   1709: 'Spare_Fault_1709', class No Acknowledgement, trigger "DB302_HMI_Faults_Carrier26_Faults_2" bit 12
   1710: 'Spare_Fault_1710', class No Acknowledgement, trigger "DB302_HMI_Faults_Carrier26_Faults_2" bit 13
   1711: 'Spare_Fault_1711', class No Acknowledgement, trigger "DB302_HMI_Faults_Carrier26_Faults_2" bit 14
   1712: 'Spare_Fault_1712', class No Acknowledgement, trigger "DB302_HMI_Faults_Carrier26_Faults_2" bit 15
   1713: 'Spare_Fault_1713', class No Acknowledgement, trigger "DB302_HMI_Faults_Carrier26_Faults_3" bit 0
   1714: 'Spare_Fault_1714', class No Acknowledgement, trigger "DB302_HMI_Faults_Carrier26_Faults_3" bit 1
   1715: 'Spare_Fault_1715', class No Acknowledgement, trigger "DB302_HMI_Faults_Carrier26_Faults_3" bit 2
   1716: 'Spare_Fault_1716', class No Acknowledgement, trigger "DB302_HMI_Faults_Carrier26_Faults_3" bit 3
   1717: 'Spare_Fault_1717', class No Acknowledgement, trigger "DB302_HMI_Faults_Carrier26_Faults_3" bit 4
   1718: 'Spare_Fault_1718', class No Acknowledgement, trigger "DB302_HMI_Faults_Carrier26_Faults_3" bit 5
   1719: 'Spare_Fault_1719', class No Acknowledgement, trigger "DB302_HMI_Faults_Carrier26_Faults_3" bit 6
   1720: 'Spare_Fault_1720', class No Acknowledgement, trigger "DB302_HMI_Faults_Carrier26_Faults_3" bit 7
   1721: 'Spare_Fault_1721', class No Acknowledgement, trigger "DB302_HMI_Faults_Carrier26_Faults_3" bit 8
   1722: 'Spare_Fault_1722', class No Acknowledgement, trigger "DB302_HMI_Faults_Carrier26_Faults_3" bit 9
   1723: 'Spare_Fault_1723', class No Acknowledgement, trigger "DB302_HMI_Faults_Carrier26_Faults_3" bit 10
   1724: 'Spare_Fault_1724', class No Acknowledgement, trigger "DB302_HMI_Faults_Carrier26_Faults_3" bit 11
   1725: 'Spare_Fault_1725', class No Acknowledgement, trigger "DB302_HMI_Faults_Carrier26_Faults_3" bit 12
   1726: 'Spare_Fault_1726', class No Acknowledgement, trigger "DB302_HMI_Faults_Carrier26_Faults_3" bit 13
   1727: 'Spare_Fault_1727', class No Acknowledgement, trigger "DB302_HMI_Faults_Carrier26_Faults_3" bit 14
   1728: 'Spare_Fault_1728', class No Acknowledgement, trigger "DB302_HMI_Faults_Carrier26_Faults_3" bit 15
   1729: 'Carrier 27 Disconnect Open Power Fault DI11.0', class No Acknowledgement, trigger "DB302_HMI_Faults_Carrier27_Faults_0" bit 0
   1730: 'Carrier 27 Drive Profinet Comm Fault', class No Acknowledgement, trigger "DB302_HMI_Faults_Carrier27_Faults_0" bit 1
   1731: 'Carrier 27 Production Stop Not Reset', class No Acknowledgement, trigger "DB302_HMI_Faults_Carrier27_Faults_0" bit 2
   1732: 'Carrier 27 CB02122 Tripped', class No Acknowledgement, trigger "DB302_HMI_Faults_Carrier27_Faults_0" bit 3
   1733: 'Carrier 27 CB02123 Tripped', class No Acknowledgement, trigger "DB302_HMI_Faults_Carrier27_Faults_0" bit 4
   1734: 'Carrier 27 AUX1 CB Tripped', class No Acknowledgement, trigger "DB302_HMI_Faults_Carrier27_Faults_0" bit 5
   1735: 'Carrier 27 AUX2 CB Tripped', class No Acknowledgement, trigger "DB302_HMI_Faults_Carrier27_Faults_0" bit 6
   1736: 'Carrier 27 PLC Not Communicating', class No Acknowledgement, trigger "DB302_HMI_Faults_Carrier27_Faults_0" bit 7
   1737: 'Carrier 27 Safe Input Card Fault', class No Acknowledgement, trigger "DB302_HMI_Faults_Carrier27_Faults_0" bit 8
   1738: 'Carrier 27 Safe Output Card Fault', class No Acknowledgement, trigger "DB302_HMI_Faults_Carrier27_Faults_0" bit 9
   1739: 'Carrier 27 Standard Input Card Fault', class No Acknowledgement, trigger "DB302_HMI_Faults_Carrier27_Faults_0" bit 10
   1740: 'Carrier 27 Standard Output Card Fault', class No Acknowledgement, trigger "DB302_HMI_Faults_Carrier27_Faults_0" bit 11
   1741: 'Carrier 27 Encoder Position Fault', class No Acknowledgement, trigger "DB302_HMI_Faults_Carrier27_Faults_0" bit 12
   1742: 'Carrier 27 Encoder Internal Error', class No Acknowledgement, trigger "DB302_HMI_Faults_Carrier27_Faults_0" bit 13
   1743: 'Carrier 27 Encoder Comm Fault', class No Acknowledgement, trigger "DB302_HMI_Faults_Carrier27_Faults_0" bit 14
   1744: 'Carrier 27 HMI Comm Fault', class No Acknowledgement, trigger "DB302_HMI_Faults_Carrier27_Faults_0" bit 15
   1745: 'Carrier 27 Crash Detection Fault', class No Acknowledgement, trigger "DB302_HMI_Faults_Carrier27_Faults_1" bit 0
   1746: 'Carrier 27 Carrier Number Invalid', class No Acknowledgement, trigger "DB302_HMI_Faults_Carrier27_Faults_1" bit 1
   1747: 'Carrier 27 Drive: PROFINET configuration error', class No Acknowledgement, trigger "DB302_HMI_Faults_Carrier27_Faults_1" bit 2
   1748: 'Carrier 27 Drive: Error internal communications', class No Acknowledgement, trigger "DB302_HMI_Faults_Carrier27_Faults_1" bit 3
   1749: 'Carrier 27 Drive: Motor overtemperature', class No Acknowledgement, trigger "DB302_HMI_Faults_Carrier27_Faults_1" bit 4
   1750: 'Carrier 27 Drive: Motor overcurrent', class No Acknowledgement, trigger "DB302_HMI_Faults_Carrier27_Faults_1" bit 5
   1751: 'Carrier 27 Drive: Infeed or power unit not ready', class No Acknowledgement, trigger "DB302_HMI_Faults_Carrier27_Faults_1" bit 6
   1752: 'Carrier 27 Drive: Short-circuit/ground fault detected', class No Acknowledgement, trigger "DB302_HMI_Faults_Carrier27_Faults_1" bit 7
   1753: 'Carrier 27 Drive: PROFINET Setpoint timeout', class No Acknowledgement, trigger "DB302_HMI_Faults_Carrier27_Faults_1" bit 8
   1754: 'Carrier 27 Power unit: Overcurrent', class No Acknowledgement, trigger "DB302_HMI_Faults_Carrier27_Faults_1" bit 9
   1755: 'Carrier 27 Power unit: DC link voltage overvoltage', class No Acknowledgement, trigger "DB302_HMI_Faults_Carrier27_Faults_1" bit 10
   1756: 'Carrier 27 Power unit: DC link voltage undervoltage', class No Acknowledgement, trigger "DB302_HMI_Faults_Carrier27_Faults_1" bit 11
   1757: 'Carrier 27 Power unit: Line phase failure in main circuit', class No Acknowledgement, trigger "DB302_HMI_Faults_Carrier27_Faults_1" bit 12
   1758: 'Carrier 27 Power unit: Phase failure motor cable', class No Acknowledgement, trigger "DB302_HMI_Faults_Carrier27_Faults_1" bit 13
   1759: 'Carrier 27 Power unit: Ground fault', class No Acknowledgement, trigger "DB302_HMI_Faults_Carrier27_Faults_1" bit 14
   1760: 'Spare_Fault_1760', class No Acknowledgement, trigger "DB302_HMI_Faults_Carrier27_Faults_1" bit 15
   1761: 'Carrier 27 Motion Off Fault', class No Acknowledgement, trigger "DB302_HMI_Faults_Carrier27_Faults_2" bit 0
   1762: 'Carrier 27 Motion On Fault', class No Acknowledgement, trigger "DB302_HMI_Faults_Carrier27_Faults_2" bit 1
   1763: 'Carrier 27 Spacing Fault', class No Acknowledgement, trigger "DB302_HMI_Faults_Carrier27_Faults_2" bit 2
   1764: 'Carrier 27 Duplicate Carrier Number Fault', class No Acknowledgement, trigger "DB302_HMI_Faults_Carrier27_Faults_2" bit 3
   1765: 'Spare_Fault_1765', class No Acknowledgement, trigger "DB302_HMI_Faults_Carrier27_Faults_2" bit 4
   1766: 'Spare_Fault_1766', class No Acknowledgement, trigger "DB302_HMI_Faults_Carrier27_Faults_2" bit 5
   1767: 'Spare_Fault_1767', class No Acknowledgement, trigger "DB302_HMI_Faults_Carrier27_Faults_2" bit 6
   1768: 'Spare_Fault_1768', class No Acknowledgement, trigger "DB302_HMI_Faults_Carrier27_Faults_2" bit 7
   1769: 'Spare_Fault_1769', class No Acknowledgement, trigger "DB302_HMI_Faults_Carrier27_Faults_2" bit 8
   1770: 'Spare_Fault_1770', class No Acknowledgement, trigger "DB302_HMI_Faults_Carrier27_Faults_2" bit 9
   1771: 'Spare_Fault_1771', class No Acknowledgement, trigger "DB302_HMI_Faults_Carrier27_Faults_2" bit 10
   1772: 'Spare_Fault_1772', class No Acknowledgement, trigger "DB302_HMI_Faults_Carrier27_Faults_2" bit 11
   1773: 'Spare_Fault_1773', class No Acknowledgement, trigger "DB302_HMI_Faults_Carrier27_Faults_2" bit 12
   1774: 'Spare_Fault_1774', class No Acknowledgement, trigger "DB302_HMI_Faults_Carrier27_Faults_2" bit 13
   1775: 'Spare_Fault_1775', class No Acknowledgement, trigger "DB302_HMI_Faults_Carrier27_Faults_2" bit 14
   1776: 'Spare_Fault_1776', class No Acknowledgement, trigger "DB302_HMI_Faults_Carrier27_Faults_2" bit 15
   1777: 'Spare_Fault_1777', class No Acknowledgement, trigger "DB302_HMI_Faults_Carrier27_Faults_3" bit 0
   1778: 'Spare_Fault_1778', class No Acknowledgement, trigger "DB302_HMI_Faults_Carrier27_Faults_3" bit 1
   1779: 'Spare_Fault_1779', class No Acknowledgement, trigger "DB302_HMI_Faults_Carrier27_Faults_3" bit 2
   1780: 'Spare_Fault_1780', class No Acknowledgement, trigger "DB302_HMI_Faults_Carrier27_Faults_3" bit 3
   1781: 'Spare_Fault_1781', class No Acknowledgement, trigger "DB302_HMI_Faults_Carrier27_Faults_3" bit 4
   1782: 'Spare_Fault_1782', class No Acknowledgement, trigger "DB302_HMI_Faults_Carrier27_Faults_3" bit 5
   1783: 'Spare_Fault_1783', class No Acknowledgement, trigger "DB302_HMI_Faults_Carrier27_Faults_3" bit 6
   1784: 'Spare_Fault_1784', class No Acknowledgement, trigger "DB302_HMI_Faults_Carrier27_Faults_3" bit 7
   1785: 'Spare_Fault_1785', class No Acknowledgement, trigger "DB302_HMI_Faults_Carrier27_Faults_3" bit 8
   1786: 'Spare_Fault_1786', class No Acknowledgement, trigger "DB302_HMI_Faults_Carrier27_Faults_3" bit 9
   1787: 'Spare_Fault_1787', class No Acknowledgement, trigger "DB302_HMI_Faults_Carrier27_Faults_3" bit 10
   1788: 'Spare_Fault_1788', class No Acknowledgement, trigger "DB302_HMI_Faults_Carrier27_Faults_3" bit 11
   1789: 'Spare_Fault_1789', class No Acknowledgement, trigger "DB302_HMI_Faults_Carrier27_Faults_3" bit 12
   1790: 'Spare_Fault_1790', class No Acknowledgement, trigger "DB302_HMI_Faults_Carrier27_Faults_3" bit 13
   1791: 'Spare_Fault_1791', class No Acknowledgement, trigger "DB302_HMI_Faults_Carrier27_Faults_3" bit 14
   1792: 'Spare_Fault_1792', class No Acknowledgement, trigger "DB302_HMI_Faults_Carrier27_Faults_3" bit 15
   1793: 'Carrier 28 Disconnect Open Power Fault DI11.0', class No Acknowledgement, trigger "DB302_HMI_Faults_Carrier28_Faults_0" bit 0
   1794: 'Carrier 28 Drive Profinet Comm Fault', class No Acknowledgement, trigger "DB302_HMI_Faults_Carrier28_Faults_0" bit 1
   1795: 'Carrier 28 Production Stop Not Reset', class No Acknowledgement, trigger "DB302_HMI_Faults_Carrier28_Faults_0" bit 2
   1796: 'Carrier 28 CB02122 Tripped', class No Acknowledgement, trigger "DB302_HMI_Faults_Carrier28_Faults_0" bit 3
   1797: 'Carrier 28 CB02123 Tripped', class No Acknowledgement, trigger "DB302_HMI_Faults_Carrier28_Faults_0" bit 4
   1798: 'Carrier 28 AUX1 CB Tripped', class No Acknowledgement, trigger "DB302_HMI_Faults_Carrier28_Faults_0" bit 5
   1799: 'Carrier 28 AUX2 CB Tripped', class No Acknowledgement, trigger "DB302_HMI_Faults_Carrier28_Faults_0" bit 6
   1800: 'Carrier 28 PLC Not Communicating', class No Acknowledgement, trigger "DB302_HMI_Faults_Carrier28_Faults_0" bit 7
   1801: 'Carrier 28 Safe Input Card Fault', class No Acknowledgement, trigger "DB302_HMI_Faults_Carrier28_Faults_0" bit 8
   1802: 'Carrier 28 Safe Output Card Fault', class No Acknowledgement, trigger "DB302_HMI_Faults_Carrier28_Faults_0" bit 9
   1803: 'Carrier 28 Standard Input Card Fault', class No Acknowledgement, trigger "DB302_HMI_Faults_Carrier28_Faults_0" bit 10
   1804: 'Carrier 28 Standard Output Card Fault', class No Acknowledgement, trigger "DB302_HMI_Faults_Carrier28_Faults_0" bit 11
   1805: 'Carrier 28 Encoder Position Fault', class No Acknowledgement, trigger "DB302_HMI_Faults_Carrier28_Faults_0" bit 12
   1806: 'Carrier 28 Encoder Internal Error', class No Acknowledgement, trigger "DB302_HMI_Faults_Carrier28_Faults_0" bit 13
   1807: 'Carrier 28 Encoder Comm Fault', class No Acknowledgement, trigger "DB302_HMI_Faults_Carrier28_Faults_0" bit 14
   1808: 'Carrier 28 HMI Comm Fault', class No Acknowledgement, trigger "DB302_HMI_Faults_Carrier28_Faults_0" bit 15
   1809: 'Carrier 28 Crash Detection Fault', class No Acknowledgement, trigger "DB302_HMI_Faults_Carrier28_Faults_1" bit 0
   1810: 'Carrier 28 Carrier Number Invalid', class No Acknowledgement, trigger "DB302_HMI_Faults_Carrier28_Faults_1" bit 1
   1811: 'Carrier 28 Drive: PROFINET configuration error', class No Acknowledgement, trigger "DB302_HMI_Faults_Carrier28_Faults_1" bit 2
   1812: 'Carrier 28 Drive: Error internal communications', class No Acknowledgement, trigger "DB302_HMI_Faults_Carrier28_Faults_1" bit 3
   1813: 'Carrier 28 Drive: Motor overtemperature', class No Acknowledgement, trigger "DB302_HMI_Faults_Carrier28_Faults_1" bit 4
   1814: 'Carrier 28 Drive: Motor overcurrent', class No Acknowledgement, trigger "DB302_HMI_Faults_Carrier28_Faults_1" bit 5
   1815: 'Carrier 28 Drive: Infeed or power unit not ready', class No Acknowledgement, trigger "DB302_HMI_Faults_Carrier28_Faults_1" bit 6
   1816: 'Carrier 28 Drive: Short-circuit/ground fault detected', class No Acknowledgement, trigger "DB302_HMI_Faults_Carrier28_Faults_1" bit 7
   1817: 'Carrier 28 Drive: PROFINET Setpoint timeout', class No Acknowledgement, trigger "DB302_HMI_Faults_Carrier28_Faults_1" bit 8
   1818: 'Carrier 28 Power unit: Overcurrent', class No Acknowledgement, trigger "DB302_HMI_Faults_Carrier28_Faults_1" bit 9
   1819: 'Carrier 28 Power unit: DC link voltage overvoltage', class No Acknowledgement, trigger "DB302_HMI_Faults_Carrier28_Faults_1" bit 10
   1820: 'Carrier 28 Power unit: DC link voltage undervoltage', class No Acknowledgement, trigger "DB302_HMI_Faults_Carrier28_Faults_1" bit 11
   1821: 'Carrier 28 Power unit: Line phase failure in main circuit', class No Acknowledgement, trigger "DB302_HMI_Faults_Carrier28_Faults_1" bit 12
   1822: 'Carrier 28 Power unit: Phase failure motor cable', class No Acknowledgement, trigger "DB302_HMI_Faults_Carrier28_Faults_1" bit 13
   1823: 'Carrier 28 Power unit: Ground fault', class No Acknowledgement, trigger "DB302_HMI_Faults_Carrier28_Faults_1" bit 14
   1824: 'Spare_Fault_1824', class No Acknowledgement, trigger "DB302_HMI_Faults_Carrier28_Faults_1" bit 15
   1825: 'Carrier 28 Motion Off Fault', class No Acknowledgement, trigger "DB302_HMI_Faults_Carrier28_Faults_2" bit 0
   1826: 'Carrier 28 Motion On Fault', class No Acknowledgement, trigger "DB302_HMI_Faults_Carrier28_Faults_2" bit 1
   1827: 'Carrier 28 Spacing Fault', class No Acknowledgement, trigger "DB302_HMI_Faults_Carrier28_Faults_2" bit 2
   1828: 'Carrier 28 Duplicate Carrier Number Fault', class No Acknowledgement, trigger "DB302_HMI_Faults_Carrier28_Faults_2" bit 3
   1829: 'Spare_Fault_1829', class No Acknowledgement, trigger "DB302_HMI_Faults_Carrier28_Faults_2" bit 4
   1830: 'Spare_Fault_1830', class No Acknowledgement, trigger "DB302_HMI_Faults_Carrier28_Faults_2" bit 5
   1831: 'Spare_Fault_1831', class No Acknowledgement, trigger "DB302_HMI_Faults_Carrier28_Faults_2" bit 6
   1832: 'Spare_Fault_1832', class No Acknowledgement, trigger "DB302_HMI_Faults_Carrier28_Faults_2" bit 7
   1833: 'Spare_Fault_1833', class No Acknowledgement, trigger "DB302_HMI_Faults_Carrier28_Faults_2" bit 8
   1834: 'Spare_Fault_1834', class No Acknowledgement, trigger "DB302_HMI_Faults_Carrier28_Faults_2" bit 9
   1835: 'Spare_Fault_1835', class No Acknowledgement, trigger "DB302_HMI_Faults_Carrier28_Faults_2" bit 10
   1836: 'Spare_Fault_1836', class No Acknowledgement, trigger "DB302_HMI_Faults_Carrier28_Faults_2" bit 11
   1837: 'Spare_Fault_1837', class No Acknowledgement, trigger "DB302_HMI_Faults_Carrier28_Faults_2" bit 12
   1838: 'Spare_Fault_1838', class No Acknowledgement, trigger "DB302_HMI_Faults_Carrier28_Faults_2" bit 13
   1839: 'Spare_Fault_1839', class No Acknowledgement, trigger "DB302_HMI_Faults_Carrier28_Faults_2" bit 14
   1840: 'Spare_Fault_1840', class No Acknowledgement, trigger "DB302_HMI_Faults_Carrier28_Faults_2" bit 15
   1841: 'Spare_Fault_1841', class No Acknowledgement, trigger "DB302_HMI_Faults_Carrier28_Faults_3" bit 0
   1842: 'Spare_Fault_1842', class No Acknowledgement, trigger "DB302_HMI_Faults_Carrier28_Faults_3" bit 1
   1843: 'Spare_Fault_1843', class No Acknowledgement, trigger "DB302_HMI_Faults_Carrier28_Faults_3" bit 2
   1844: 'Spare_Fault_1844', class No Acknowledgement, trigger "DB302_HMI_Faults_Carrier28_Faults_3" bit 3
   1845: 'Spare_Fault_1845', class No Acknowledgement, trigger "DB302_HMI_Faults_Carrier28_Faults_3" bit 4
   1846: 'Spare_Fault_1846', class No Acknowledgement, trigger "DB302_HMI_Faults_Carrier28_Faults_3" bit 5
   1847: 'Spare_Fault_1847', class No Acknowledgement, trigger "DB302_HMI_Faults_Carrier28_Faults_3" bit 6
   1848: 'Spare_Fault_1848', class No Acknowledgement, trigger "DB302_HMI_Faults_Carrier28_Faults_3" bit 7
   1849: 'Spare_Fault_1849', class No Acknowledgement, trigger "DB302_HMI_Faults_Carrier28_Faults_3" bit 8
   1850: 'Spare_Fault_1850', class No Acknowledgement, trigger "DB302_HMI_Faults_Carrier28_Faults_3" bit 9
   1851: 'Spare_Fault_1851', class No Acknowledgement, trigger "DB302_HMI_Faults_Carrier28_Faults_3" bit 10
   1852: 'Spare_Fault_1852', class No Acknowledgement, trigger "DB302_HMI_Faults_Carrier28_Faults_3" bit 11
   1853: 'Spare_Fault_1853', class No Acknowledgement, trigger "DB302_HMI_Faults_Carrier28_Faults_3" bit 12
   1854: 'Spare_Fault_1854', class No Acknowledgement, trigger "DB302_HMI_Faults_Carrier28_Faults_3" bit 13
   1855: 'Spare_Fault_1855', class No Acknowledgement, trigger "DB302_HMI_Faults_Carrier28_Faults_3" bit 14
   1856: 'Spare_Fault_1856', class No Acknowledgement, trigger "DB302_HMI_Faults_Carrier28_Faults_3" bit 15
   1857: 'Carrier 29 Disconnect Open Power Fault DI11.0', class No Acknowledgement, trigger "DB302_HMI_Faults_Carrier29_Faults_0" bit 0
   1858: 'Carrier 29 Drive Profinet Comm Fault', class No Acknowledgement, trigger "DB302_HMI_Faults_Carrier29_Faults_0" bit 1
   1859: 'Carrier 29 Production Stop Not Reset', class No Acknowledgement, trigger "DB302_HMI_Faults_Carrier29_Faults_0" bit 2
   1860: 'Carrier 29 CB02122 Tripped', class No Acknowledgement, trigger "DB302_HMI_Faults_Carrier29_Faults_0" bit 3
   1861: 'Carrier 29 CB02123 Tripped', class No Acknowledgement, trigger "DB302_HMI_Faults_Carrier29_Faults_0" bit 4
   1862: 'Carrier 29 AUX1 CB Tripped', class No Acknowledgement, trigger "DB302_HMI_Faults_Carrier29_Faults_0" bit 5
   1863: 'Carrier 29 AUX2 CB Tripped', class No Acknowledgement, trigger "DB302_HMI_Faults_Carrier29_Faults_0" bit 6
   1864: 'Carrier 29 PLC Not Communicating', class No Acknowledgement, trigger "DB302_HMI_Faults_Carrier29_Faults_0" bit 7
   1865: 'Carrier 29 Safe Input Card Fault', class No Acknowledgement, trigger "DB302_HMI_Faults_Carrier29_Faults_0" bit 8
   1866: 'Carrier 29 Safe Output Card Fault', class No Acknowledgement, trigger "DB302_HMI_Faults_Carrier29_Faults_0" bit 9
   1867: 'Carrier 29 Standard Input Card Fault', class No Acknowledgement, trigger "DB302_HMI_Faults_Carrier29_Faults_0" bit 10
   1868: 'Carrier 29 Standard Output Card Fault', class No Acknowledgement, trigger "DB302_HMI_Faults_Carrier29_Faults_0" bit 11
   1869: 'Carrier 29 Encoder Position Fault', class No Acknowledgement, trigger "DB302_HMI_Faults_Carrier29_Faults_0" bit 12
   1870: 'Carrier 29 Encoder Internal Error', class No Acknowledgement, trigger "DB302_HMI_Faults_Carrier29_Faults_0" bit 13
   1871: 'Carrier 29 Encoder Comm Fault', class No Acknowledgement, trigger "DB302_HMI_Faults_Carrier29_Faults_0" bit 14
   1872: 'Carrier 29 HMI Comm Fault', class No Acknowledgement, trigger "DB302_HMI_Faults_Carrier29_Faults_0" bit 15
   1873: 'Carrier 29 Crash Detection Fault', class No Acknowledgement, trigger "DB302_HMI_Faults_Carrier29_Faults_1" bit 0
   1874: 'Carrier 29 Carrier Number Invalid', class No Acknowledgement, trigger "DB302_HMI_Faults_Carrier29_Faults_1" bit 1
   1875: 'Carrier 29 Drive: PROFINET configuration error', class No Acknowledgement, trigger "DB302_HMI_Faults_Carrier29_Faults_1" bit 2
   1876: 'Carrier 29 Drive: Error internal communications', class No Acknowledgement, trigger "DB302_HMI_Faults_Carrier29_Faults_1" bit 3
   1877: 'Carrier 29 Drive: Motor overtemperature', class No Acknowledgement, trigger "DB302_HMI_Faults_Carrier29_Faults_1" bit 4
   1878: 'Carrier 29 Drive: Motor overcurrent', class No Acknowledgement, trigger "DB302_HMI_Faults_Carrier29_Faults_1" bit 5
   1879: 'Carrier 29 Drive: Infeed or power unit not ready', class No Acknowledgement, trigger "DB302_HMI_Faults_Carrier29_Faults_1" bit 6
   1880: 'Carrier 29 Drive: Short-circuit/ground fault detected', class No Acknowledgement, trigger "DB302_HMI_Faults_Carrier29_Faults_1" bit 7
   1881: 'Carrier 29 Drive: PROFINET Setpoint timeout', class No Acknowledgement, trigger "DB302_HMI_Faults_Carrier29_Faults_1" bit 8
   1882: 'Carrier 29 Power unit: Overcurrent', class No Acknowledgement, trigger "DB302_HMI_Faults_Carrier29_Faults_1" bit 9
   1883: 'Carrier 29 Power unit: DC link voltage overvoltage', class No Acknowledgement, trigger "DB302_HMI_Faults_Carrier29_Faults_1" bit 10
   1884: 'Carrier 29 Power unit: DC link voltage undervoltage', class No Acknowledgement, trigger "DB302_HMI_Faults_Carrier29_Faults_1" bit 11
   1885: 'Carrier 29 Power unit: Line phase failure in main circuit', class No Acknowledgement, trigger "DB302_HMI_Faults_Carrier29_Faults_1" bit 12
   1886: 'Carrier 29 Power unit: Phase failure motor cable', class No Acknowledgement, trigger "DB302_HMI_Faults_Carrier29_Faults_1" bit 13
   1887: 'Carrier 29 Power unit: Ground fault', class No Acknowledgement, trigger "DB302_HMI_Faults_Carrier29_Faults_1" bit 14
   1888: 'Spare_Fault_1888', class No Acknowledgement, trigger "DB302_HMI_Faults_Carrier29_Faults_1" bit 15
   1889: 'Carrier 29 Motion Off Fault', class No Acknowledgement, trigger "DB302_HMI_Faults_Carrier29_Faults_2" bit 0
   1890: 'Carrier 29 Motion On Fault', class No Acknowledgement, trigger "DB302_HMI_Faults_Carrier29_Faults_2" bit 1
   1891: 'Carrier 29 Spacing Fault', class No Acknowledgement, trigger "DB302_HMI_Faults_Carrier29_Faults_2" bit 2
   1892: 'Carrier 29 Duplicate Carrier Number Fault', class No Acknowledgement, trigger "DB302_HMI_Faults_Carrier29_Faults_2" bit 3
   1893: 'Spare_Fault_1893', class No Acknowledgement, trigger "DB302_HMI_Faults_Carrier29_Faults_2" bit 4
   1894: 'Spare_Fault_1894', class No Acknowledgement, trigger "DB302_HMI_Faults_Carrier29_Faults_2" bit 5
   1895: 'Spare_Fault_1895', class No Acknowledgement, trigger "DB302_HMI_Faults_Carrier29_Faults_2" bit 6
   1896: 'Spare_Fault_1896', class No Acknowledgement, trigger "DB302_HMI_Faults_Carrier29_Faults_2" bit 7
   1897: 'Spare_Fault_1897', class No Acknowledgement, trigger "DB302_HMI_Faults_Carrier29_Faults_2" bit 8
   1898: 'Spare_Fault_1898', class No Acknowledgement, trigger "DB302_HMI_Faults_Carrier29_Faults_2" bit 9
   1899: 'Spare_Fault_1899', class No Acknowledgement, trigger "DB302_HMI_Faults_Carrier29_Faults_2" bit 10
   1900: 'Spare_Fault_1900', class No Acknowledgement, trigger "DB302_HMI_Faults_Carrier29_Faults_2" bit 11
   1901: 'Spare_Fault_1901', class No Acknowledgement, trigger "DB302_HMI_Faults_Carrier29_Faults_2" bit 12
   1902: 'Spare_Fault_1902', class No Acknowledgement, trigger "DB302_HMI_Faults_Carrier29_Faults_2" bit 13
   1903: 'Spare_Fault_1903', class No Acknowledgement, trigger "DB302_HMI_Faults_Carrier29_Faults_2" bit 14
   1904: 'Spare_Fault_1904', class No Acknowledgement, trigger "DB302_HMI_Faults_Carrier29_Faults_2" bit 15
   1905: 'Spare_Fault_1905', class No Acknowledgement, trigger "DB302_HMI_Faults_Carrier29_Faults_3" bit 0
   1906: 'Spare_Fault_1906', class No Acknowledgement, trigger "DB302_HMI_Faults_Carrier29_Faults_3" bit 1
   1907: 'Spare_Fault_1907', class No Acknowledgement, trigger "DB302_HMI_Faults_Carrier29_Faults_3" bit 2
   1908: 'Spare_Fault_1908', class No Acknowledgement, trigger "DB302_HMI_Faults_Carrier29_Faults_3" bit 3
   1909: 'Spare_Fault_1909', class No Acknowledgement, trigger "DB302_HMI_Faults_Carrier29_Faults_3" bit 4
   1910: 'Spare_Fault_1910', class No Acknowledgement, trigger "DB302_HMI_Faults_Carrier29_Faults_3" bit 5
   1911: 'Spare_Fault_1911', class No Acknowledgement, trigger "DB302_HMI_Faults_Carrier29_Faults_3" bit 6
   1912: 'Spare_Fault_1912', class No Acknowledgement, trigger "DB302_HMI_Faults_Carrier29_Faults_3" bit 7
   1913: 'Spare_Fault_1913', class No Acknowledgement, trigger "DB302_HMI_Faults_Carrier29_Faults_3" bit 8
   1914: 'Spare_Fault_1914', class No Acknowledgement, trigger "DB302_HMI_Faults_Carrier29_Faults_3" bit 9
   1915: 'Spare_Fault_1915', class No Acknowledgement, trigger "DB302_HMI_Faults_Carrier29_Faults_3" bit 10
   1916: 'Spare_Fault_1916', class No Acknowledgement, trigger "DB302_HMI_Faults_Carrier29_Faults_3" bit 11
   1917: 'Spare_Fault_1917', class No Acknowledgement, trigger "DB302_HMI_Faults_Carrier29_Faults_3" bit 12
   1918: 'Spare_Fault_1918', class No Acknowledgement, trigger "DB302_HMI_Faults_Carrier29_Faults_3" bit 13
   1919: 'Spare_Fault_1919', class No Acknowledgement, trigger "DB302_HMI_Faults_Carrier29_Faults_3" bit 14
   1920: 'Spare_Fault_1920', class No Acknowledgement, trigger "DB302_HMI_Faults_Carrier29_Faults_3" bit 15
   1921: 'Carrier 30 Disconnect Open Power Fault DI11.0', class No Acknowledgement, trigger "DB302_HMI_Faults_Carrier30_Faults_0" bit 0
   1922: 'Carrier 30 Drive Profinet Comm Fault', class No Acknowledgement, trigger "DB302_HMI_Faults_Carrier30_Faults_0" bit 1
   1923: 'Carrier 30 Production Stop Not Reset', class No Acknowledgement, trigger "DB302_HMI_Faults_Carrier30_Faults_0" bit 2
   1924: 'Carrier 30 CB02122 Tripped', class No Acknowledgement, trigger "DB302_HMI_Faults_Carrier30_Faults_0" bit 3
   1925: 'Carrier 30 CB02123 Tripped', class No Acknowledgement, trigger "DB302_HMI_Faults_Carrier30_Faults_0" bit 4
   1926: 'Carrier 30 AUX1 CB Tripped', class No Acknowledgement, trigger "DB302_HMI_Faults_Carrier30_Faults_0" bit 5
   1927: 'Carrier 30 AUX2 CB Tripped', class No Acknowledgement, trigger "DB302_HMI_Faults_Carrier30_Faults_0" bit 6
   1928: 'Carrier 30 PLC Not Communicating', class No Acknowledgement, trigger "DB302_HMI_Faults_Carrier30_Faults_0" bit 7
   1929: 'Carrier 30 Safe Input Card Fault', class No Acknowledgement, trigger "DB302_HMI_Faults_Carrier30_Faults_0" bit 8
   1930: 'Carrier 30 Safe Output Card Fault', class No Acknowledgement, trigger "DB302_HMI_Faults_Carrier30_Faults_0" bit 9
   1931: 'Carrier 30 Standard Input Card Fault', class No Acknowledgement, trigger "DB302_HMI_Faults_Carrier30_Faults_0" bit 10
   1932: 'Carrier 30 Standard Output Card Fault', class No Acknowledgement, trigger "DB302_HMI_Faults_Carrier30_Faults_0" bit 11
   1933: 'Carrier 30 Encoder Position Fault', class No Acknowledgement, trigger "DB302_HMI_Faults_Carrier30_Faults_0" bit 12
   1934: 'Carrier 30 Encoder Internal Error', class No Acknowledgement, trigger "DB302_HMI_Faults_Carrier30_Faults_0" bit 13
   1935: 'Carrier 30 Encoder Comm Fault', class No Acknowledgement, trigger "DB302_HMI_Faults_Carrier30_Faults_0" bit 14
   1936: 'Carrier 30 HMI Comm Fault', class No Acknowledgement, trigger "DB302_HMI_Faults_Carrier30_Faults_0" bit 15
   1937: 'Carrier 30 Crash Detection Fault', class No Acknowledgement, trigger "DB302_HMI_Faults_Carrier30_Faults_1" bit 0
   1938: 'Carrier 30 Carrier Number Invalid', class No Acknowledgement, trigger "DB302_HMI_Faults_Carrier30_Faults_1" bit 1
   1939: 'Carrier 30 Drive: PROFINET configuration error', class No Acknowledgement, trigger "DB302_HMI_Faults_Carrier30_Faults_1" bit 2
   1940: 'Carrier 30 Drive: Error internal communications', class No Acknowledgement, trigger "DB302_HMI_Faults_Carrier30_Faults_1" bit 3
   1941: 'Carrier 30 Drive: Motor overtemperature', class No Acknowledgement, trigger "DB302_HMI_Faults_Carrier30_Faults_1" bit 4
   1942: 'Carrier 30 Drive: Motor overcurrent', class No Acknowledgement, trigger "DB302_HMI_Faults_Carrier30_Faults_1" bit 5
   1943: 'Carrier 30 Drive: Infeed or power unit not ready', class No Acknowledgement, trigger "DB302_HMI_Faults_Carrier30_Faults_1" bit 6
   1944: 'Carrier 30 Drive: Short-circuit/ground fault detected', class No Acknowledgement, trigger "DB302_HMI_Faults_Carrier30_Faults_1" bit 7
   1945: 'Carrier 30 Drive: PROFINET Setpoint timeout', class No Acknowledgement, trigger "DB302_HMI_Faults_Carrier30_Faults_1" bit 8
   1946: 'Carrier 30 Power unit: Overcurrent', class No Acknowledgement, trigger "DB302_HMI_Faults_Carrier30_Faults_1" bit 9
   1947: 'Carrier 30 Power unit: DC link voltage overvoltage', class No Acknowledgement, trigger "DB302_HMI_Faults_Carrier30_Faults_1" bit 10
   1948: 'Carrier 30 Power unit: DC link voltage undervoltage', class No Acknowledgement, trigger "DB302_HMI_Faults_Carrier30_Faults_1" bit 11
   1949: 'Carrier 30 Power unit: Line phase failure in main circuit', class No Acknowledgement, trigger "DB302_HMI_Faults_Carrier30_Faults_1" bit 12
   1950: 'Carrier 30 Power unit: Phase failure motor cable', class No Acknowledgement, trigger "DB302_HMI_Faults_Carrier30_Faults_1" bit 13
   1951: 'Carrier 30 Power unit: Ground fault', class No Acknowledgement, trigger "DB302_HMI_Faults_Carrier30_Faults_1" bit 14
   1952: 'Spare_Fault_1952', class No Acknowledgement, trigger "DB302_HMI_Faults_Carrier30_Faults_1" bit 15
   1953: 'Carrier 30 Motion Off Fault', class No Acknowledgement, trigger "DB302_HMI_Faults_Carrier30_Faults_2" bit 0
   1954: 'Carrier 30 Motion On Fault', class No Acknowledgement, trigger "DB302_HMI_Faults_Carrier30_Faults_2" bit 1
   1955: 'Carrier 30 Spacing Fault', class No Acknowledgement, trigger "DB302_HMI_Faults_Carrier30_Faults_2" bit 2
   1956: 'Carrier 30 Duplicate Carrier Number Fault', class No Acknowledgement, trigger "DB302_HMI_Faults_Carrier30_Faults_2" bit 3
   1957: 'Spare_Fault_1957', class No Acknowledgement, trigger "DB302_HMI_Faults_Carrier30_Faults_2" bit 4
   1958: 'Spare_Fault_1958', class No Acknowledgement, trigger "DB302_HMI_Faults_Carrier30_Faults_2" bit 5
   1959: 'Spare_Fault_1959', class No Acknowledgement, trigger "DB302_HMI_Faults_Carrier30_Faults_2" bit 6
   1960: 'Spare_Fault_1960', class No Acknowledgement, trigger "DB302_HMI_Faults_Carrier30_Faults_2" bit 7
   1961: 'Spare_Fault_1961', class No Acknowledgement, trigger "DB302_HMI_Faults_Carrier30_Faults_2" bit 8
   1962: 'Spare_Fault_1962', class No Acknowledgement, trigger "DB302_HMI_Faults_Carrier30_Faults_2" bit 9
   1963: 'Spare_Fault_1963', class No Acknowledgement, trigger "DB302_HMI_Faults_Carrier30_Faults_2" bit 10
   1964: 'Spare_Fault_1964', class No Acknowledgement, trigger "DB302_HMI_Faults_Carrier30_Faults_2" bit 11
   1965: 'Spare_Fault_1965', class No Acknowledgement, trigger "DB302_HMI_Faults_Carrier30_Faults_2" bit 12
   1966: 'Spare_Fault_1966', class No Acknowledgement, trigger "DB302_HMI_Faults_Carrier30_Faults_2" bit 13
   1967: 'Spare_Fault_1967', class No Acknowledgement, trigger "DB302_HMI_Faults_Carrier30_Faults_2" bit 14
   1968: 'Spare_Fault_1968', class No Acknowledgement, trigger "DB302_HMI_Faults_Carrier30_Faults_2" bit 15
   1969: 'Spare_Fault_1969', class No Acknowledgement, trigger "DB302_HMI_Faults_Carrier30_Faults_3" bit 0
   1970: 'Spare_Fault_1970', class No Acknowledgement, trigger "DB302_HMI_Faults_Carrier30_Faults_3" bit 1
   1971: 'Spare_Fault_1971', class No Acknowledgement, trigger "DB302_HMI_Faults_Carrier30_Faults_3" bit 2
   1972: 'Spare_Fault_1972', class No Acknowledgement, trigger "DB302_HMI_Faults_Carrier30_Faults_3" bit 3
   1973: 'Spare_Fault_1973', class No Acknowledgement, trigger "DB302_HMI_Faults_Carrier30_Faults_3" bit 4
   1974: 'Spare_Fault_1974', class No Acknowledgement, trigger "DB302_HMI_Faults_Carrier30_Faults_3" bit 5
   1975: 'Spare_Fault_1975', class No Acknowledgement, trigger "DB302_HMI_Faults_Carrier30_Faults_3" bit 6
   1976: 'Spare_Fault_1976', class No Acknowledgement, trigger "DB302_HMI_Faults_Carrier30_Faults_3" bit 7
   1977: 'Spare_Fault_1977', class No Acknowledgement, trigger "DB302_HMI_Faults_Carrier30_Faults_3" bit 8
   1978: 'Spare_Fault_1978', class No Acknowledgement, trigger "DB302_HMI_Faults_Carrier30_Faults_3" bit 9
   1979: 'Spare_Fault_1979', class No Acknowledgement, trigger "DB302_HMI_Faults_Carrier30_Faults_3" bit 10
   1980: 'Spare_Fault_1980', class No Acknowledgement, trigger "DB302_HMI_Faults_Carrier30_Faults_3" bit 11
   1981: 'Spare_Fault_1981', class No Acknowledgement, trigger "DB302_HMI_Faults_Carrier30_Faults_3" bit 12
   1982: 'Spare_Fault_1982', class No Acknowledgement, trigger "DB302_HMI_Faults_Carrier30_Faults_3" bit 13
   1983: 'Spare_Fault_1983', class No Acknowledgement, trigger "DB302_HMI_Faults_Carrier30_Faults_3" bit 14
   1984: 'Spare_Fault_1984', class No Acknowledgement, trigger "DB302_HMI_Faults_Carrier30_Faults_3" bit 15
   1985: 'Carrier 31 Disconnect Open Power Fault DI11.0', class No Acknowledgement, trigger "DB302_HMI_Faults_Carrier31_Faults_0" bit 0
   1986: 'Carrier 31 Drive Profinet Comm Fault', class No Acknowledgement, trigger "DB302_HMI_Faults_Carrier31_Faults_0" bit 1
   1987: 'Carrier 31 Production Stop Not Reset', class No Acknowledgement, trigger "DB302_HMI_Faults_Carrier31_Faults_0" bit 2
   1988: 'Carrier 31 CB02122 Tripped', class No Acknowledgement, trigger "DB302_HMI_Faults_Carrier31_Faults_0" bit 3
   1989: 'Carrier 31 CB02123 Tripped', class No Acknowledgement, trigger "DB302_HMI_Faults_Carrier31_Faults_0" bit 4
   1990: 'Carrier 31 AUX1 CB Tripped', class No Acknowledgement, trigger "DB302_HMI_Faults_Carrier31_Faults_0" bit 5
   1991: 'Carrier 31 AUX2 CB Tripped', class No Acknowledgement, trigger "DB302_HMI_Faults_Carrier31_Faults_0" bit 6
   1992: 'Carrier 31 PLC Not Communicating', class No Acknowledgement, trigger "DB302_HMI_Faults_Carrier31_Faults_0" bit 7
   1993: 'Carrier 31 Safe Input Card Fault', class No Acknowledgement, trigger "DB302_HMI_Faults_Carrier31_Faults_0" bit 8
   1994: 'Carrier 31 Safe Output Card Fault', class No Acknowledgement, trigger "DB302_HMI_Faults_Carrier31_Faults_0" bit 9
   1995: 'Carrier 31 Standard Input Card Fault', class No Acknowledgement, trigger "DB302_HMI_Faults_Carrier31_Faults_0" bit 10
   1996: 'Carrier 31 Standard Output Card Fault', class No Acknowledgement, trigger "DB302_HMI_Faults_Carrier31_Faults_0" bit 11
   1997: 'Carrier 31 Encoder Position Fault', class No Acknowledgement, trigger "DB302_HMI_Faults_Carrier31_Faults_0" bit 12
   1998: 'Carrier 31 Encoder Internal Error', class No Acknowledgement, trigger "DB302_HMI_Faults_Carrier31_Faults_0" bit 13
   1999: 'Carrier 31 Encoder Comm Fault', class No Acknowledgement, trigger "DB302_HMI_Faults_Carrier31_Faults_0" bit 14
   2000: 'Carrier 31 HMI Comm Fault', class No Acknowledgement, trigger "DB302_HMI_Faults_Carrier31_Faults_0" bit 15
   2001: 'Carrier 31 Crash Detection Fault', class No Acknowledgement, trigger "DB302_HMI_Faults_Carrier31_Faults_1" bit 0
   2002: 'Carrier 31 Carrier Number Invalid', class No Acknowledgement, trigger "DB302_HMI_Faults_Carrier31_Faults_1" bit 1
   2003: 'Carrier 31 Drive: PROFINET configuration error', class No Acknowledgement, trigger "DB302_HMI_Faults_Carrier31_Faults_1" bit 2
   2004: 'Carrier 31 Drive: Error internal communications', class No Acknowledgement, trigger "DB302_HMI_Faults_Carrier31_Faults_1" bit 3
   2005: 'Carrier 31 Drive: Motor overtemperature', class No Acknowledgement, trigger "DB302_HMI_Faults_Carrier31_Faults_1" bit 4
   2006: 'Carrier 31 Drive: Motor overcurrent', class No Acknowledgement, trigger "DB302_HMI_Faults_Carrier31_Faults_1" bit 5
   2007: 'Carrier 31 Drive: Infeed or power unit not ready', class No Acknowledgement, trigger "DB302_HMI_Faults_Carrier31_Faults_1" bit 6
   2008: 'Carrier 31 Drive: Short-circuit/ground fault detected', class No Acknowledgement, trigger "DB302_HMI_Faults_Carrier31_Faults_1" bit 7
   2009: 'Carrier 31 Drive: PROFINET Setpoint timeout', class No Acknowledgement, trigger "DB302_HMI_Faults_Carrier31_Faults_1" bit 8
   2010: 'Carrier 31 Power unit: Overcurrent', class No Acknowledgement, trigger "DB302_HMI_Faults_Carrier31_Faults_1" bit 9
   2011: 'Carrier 31 Power unit: DC link voltage overvoltage', class No Acknowledgement, trigger "DB302_HMI_Faults_Carrier31_Faults_1" bit 10
   2012: 'Carrier 31 Power unit: DC link voltage undervoltage', class No Acknowledgement, trigger "DB302_HMI_Faults_Carrier31_Faults_1" bit 11
   2013: 'Carrier 31 Power unit: Line phase failure in main circuit', class No Acknowledgement, trigger "DB302_HMI_Faults_Carrier31_Faults_1" bit 12
   2014: 'Carrier 31 Power unit: Phase failure motor cable', class No Acknowledgement, trigger "DB302_HMI_Faults_Carrier31_Faults_1" bit 13
   2015: 'Carrier 31 Power unit: Ground fault', class No Acknowledgement, trigger "DB302_HMI_Faults_Carrier31_Faults_1" bit 14
   2016: 'Spare_Fault_2016', class No Acknowledgement, trigger "DB302_HMI_Faults_Carrier31_Faults_1" bit 15
   2017: 'Carrier 31 Motion Off Fault', class No Acknowledgement, trigger "DB302_HMI_Faults_Carrier31_Faults_2" bit 0
   2018: 'Carrier 31 Motion On Fault', class No Acknowledgement, trigger "DB302_HMI_Faults_Carrier31_Faults_2" bit 1
   2019: 'Carrier 31 Spacing Fault', class No Acknowledgement, trigger "DB302_HMI_Faults_Carrier31_Faults_2" bit 2
   2020: 'Carrier 31 Duplicate Carrier Number Fault', class No Acknowledgement, trigger "DB302_HMI_Faults_Carrier31_Faults_2" bit 3
   2021: 'Spare_Fault_2021', class No Acknowledgement, trigger "DB302_HMI_Faults_Carrier31_Faults_2" bit 4
   2022: 'Spare_Fault_2022', class No Acknowledgement, trigger "DB302_HMI_Faults_Carrier31_Faults_2" bit 5
   2023: 'Spare_Fault_2023', class No Acknowledgement, trigger "DB302_HMI_Faults_Carrier31_Faults_2" bit 6
   2024: 'Spare_Fault_2024', class No Acknowledgement, trigger "DB302_HMI_Faults_Carrier31_Faults_2" bit 7
   2025: 'Spare_Fault_2025', class No Acknowledgement, trigger "DB302_HMI_Faults_Carrier31_Faults_2" bit 8
   2026: 'Spare_Fault_2026', class No Acknowledgement, trigger "DB302_HMI_Faults_Carrier31_Faults_2" bit 9
   2027: 'Spare_Fault_2027', class No Acknowledgement, trigger "DB302_HMI_Faults_Carrier31_Faults_2" bit 10
   2028: 'Spare_Fault_2028', class No Acknowledgement, trigger "DB302_HMI_Faults_Carrier31_Faults_2" bit 11
   2029: 'Spare_Fault_2029', class No Acknowledgement, trigger "DB302_HMI_Faults_Carrier31_Faults_2" bit 12
   2030: 'Spare_Fault_2030', class No Acknowledgement, trigger "DB302_HMI_Faults_Carrier31_Faults_2" bit 13
   2031: 'Spare_Fault_2031', class No Acknowledgement, trigger "DB302_HMI_Faults_Carrier31_Faults_2" bit 14
   2032: 'Spare_Fault_2032', class No Acknowledgement, trigger "DB302_HMI_Faults_Carrier31_Faults_2" bit 15
   2033: 'Spare_Fault_2033', class No Acknowledgement, trigger "DB302_HMI_Faults_Carrier31_Faults_3" bit 0
   2034: 'Spare_Fault_2034', class No Acknowledgement, trigger "DB302_HMI_Faults_Carrier31_Faults_3" bit 1
   2035: 'Spare_Fault_2035', class No Acknowledgement, trigger "DB302_HMI_Faults_Carrier31_Faults_3" bit 2
   2036: 'Spare_Fault_2036', class No Acknowledgement, trigger "DB302_HMI_Faults_Carrier31_Faults_3" bit 3
   2037: 'Spare_Fault_2037', class No Acknowledgement, trigger "DB302_HMI_Faults_Carrier31_Faults_3" bit 4
   2038: 'Spare_Fault_2038', class No Acknowledgement, trigger "DB302_HMI_Faults_Carrier31_Faults_3" bit 5
   2039: 'Spare_Fault_2039', class No Acknowledgement, trigger "DB302_HMI_Faults_Carrier31_Faults_3" bit 6
   2040: 'Spare_Fault_2040', class No Acknowledgement, trigger "DB302_HMI_Faults_Carrier31_Faults_3" bit 7
   2041: 'Spare_Fault_2041', class No Acknowledgement, trigger "DB302_HMI_Faults_Carrier31_Faults_3" bit 8
   2042: 'Spare_Fault_2042', class No Acknowledgement, trigger "DB302_HMI_Faults_Carrier31_Faults_3" bit 9
   2043: 'Spare_Fault_2043', class No Acknowledgement, trigger "DB302_HMI_Faults_Carrier31_Faults_3" bit 10
   2044: 'Spare_Fault_2044', class No Acknowledgement, trigger "DB302_HMI_Faults_Carrier31_Faults_3" bit 11
   2045: 'Spare_Fault_2045', class No Acknowledgement, trigger "DB302_HMI_Faults_Carrier31_Faults_3" bit 12
   2046: 'Spare_Fault_2046', class No Acknowledgement, trigger "DB302_HMI_Faults_Carrier31_Faults_3" bit 13
   2047: 'Spare_Fault_2047', class No Acknowledgement, trigger "DB302_HMI_Faults_Carrier31_Faults_3" bit 14
   2048: 'Spare_Fault_2048', class No Acknowledgement, trigger "DB302_HMI_Faults_Carrier31_Faults_3" bit 15
   2049: 'Carrier 32 Disconnect Open Power Fault DI11.0', class No Acknowledgement, trigger "DB302_HMI_Faults_Carrier32_Faults_0" bit 0
   2050: 'Carrier 32 Drive Profinet Comm Fault', class No Acknowledgement, trigger "DB302_HMI_Faults_Carrier32_Faults_0" bit 1
   2051: 'Carrier 32 Production Stop Not Reset', class No Acknowledgement, trigger "DB302_HMI_Faults_Carrier32_Faults_0" bit 2
   2052: 'Carrier 32 CB02122 Tripped', class No Acknowledgement, trigger "DB302_HMI_Faults_Carrier32_Faults_0" bit 3
   2053: 'Carrier 32 CB02123 Tripped', class No Acknowledgement, trigger "DB302_HMI_Faults_Carrier32_Faults_0" bit 4
   2054: 'Carrier 32 AUX1 CB Tripped', class No Acknowledgement, trigger "DB302_HMI_Faults_Carrier32_Faults_0" bit 5
   2055: 'Carrier 32 AUX2 CB Tripped', class No Acknowledgement, trigger "DB302_HMI_Faults_Carrier32_Faults_0" bit 6
   2056: 'Carrier 32 PLC Not Communicating', class No Acknowledgement, trigger "DB302_HMI_Faults_Carrier32_Faults_0" bit 7
   2057: 'Carrier 32 Safe Input Card Fault', class No Acknowledgement, trigger "DB302_HMI_Faults_Carrier32_Faults_0" bit 8
   2058: 'Carrier 32 Safe Output Card Fault', class No Acknowledgement, trigger "DB302_HMI_Faults_Carrier32_Faults_0" bit 9
   2059: 'Carrier 32 Standard Input Card Fault', class No Acknowledgement, trigger "DB302_HMI_Faults_Carrier32_Faults_0" bit 10
   2060: 'Carrier 32 Standard Output Card Fault', class No Acknowledgement, trigger "DB302_HMI_Faults_Carrier32_Faults_0" bit 11
   2061: 'Carrier 32 Encoder Position Fault', class No Acknowledgement, trigger "DB302_HMI_Faults_Carrier32_Faults_0" bit 12
   2062: 'Carrier 32 Encoder Internal Error', class No Acknowledgement, trigger "DB302_HMI_Faults_Carrier32_Faults_0" bit 13
   2063: 'Carrier 32 Encoder Comm Fault', class No Acknowledgement, trigger "DB302_HMI_Faults_Carrier32_Faults_0" bit 14
   2064: 'Carrier 32 HMI Comm Fault', class No Acknowledgement, trigger "DB302_HMI_Faults_Carrier32_Faults_0" bit 15
   2065: 'Carrier 32 Crash Detection Fault', class No Acknowledgement, trigger "DB302_HMI_Faults_Carrier32_Faults_1" bit 0
   2066: 'Carrier 32 Carrier Number Invalid', class No Acknowledgement, trigger "DB302_HMI_Faults_Carrier32_Faults_1" bit 1
   2067: 'Carrier 32 Drive: PROFINET configuration error', class No Acknowledgement, trigger "DB302_HMI_Faults_Carrier32_Faults_1" bit 2
   2068: 'Carrier 32 Drive: Error internal communications', class No Acknowledgement, trigger "DB302_HMI_Faults_Carrier32_Faults_1" bit 3
   2069: 'Carrier 32 Drive: Motor overtemperature', class No Acknowledgement, trigger "DB302_HMI_Faults_Carrier32_Faults_1" bit 4
   2070: 'Carrier 32 Drive: Motor overcurrent', class No Acknowledgement, trigger "DB302_HMI_Faults_Carrier32_Faults_1" bit 5
   2071: 'Carrier 32 Drive: Infeed or power unit not ready', class No Acknowledgement, trigger "DB302_HMI_Faults_Carrier32_Faults_1" bit 6
   2072: 'Carrier 32 Drive: Short-circuit/ground fault detected', class No Acknowledgement, trigger "DB302_HMI_Faults_Carrier32_Faults_1" bit 7
   2073: 'Carrier 32 Drive: PROFINET Setpoint timeout', class No Acknowledgement, trigger "DB302_HMI_Faults_Carrier32_Faults_1" bit 8
   2074: 'Carrier 32 Power unit: Overcurrent', class No Acknowledgement, trigger "DB302_HMI_Faults_Carrier32_Faults_1" bit 9
   2075: 'Carrier 32 Power unit: DC link voltage overvoltage', class No Acknowledgement, trigger "DB302_HMI_Faults_Carrier32_Faults_1" bit 10
   2076: 'Carrier 32 Power unit: DC link voltage undervoltage', class No Acknowledgement, trigger "DB302_HMI_Faults_Carrier32_Faults_1" bit 11
   2077: 'Carrier 32 Power unit: Line phase failure in main circuit', class No Acknowledgement, trigger "DB302_HMI_Faults_Carrier32_Faults_1" bit 12
   2078: 'Carrier 32 Power unit: Phase failure motor cable', class No Acknowledgement, trigger "DB302_HMI_Faults_Carrier32_Faults_1" bit 13
   2079: 'Carrier 32 Power unit: Ground fault', class No Acknowledgement, trigger "DB302_HMI_Faults_Carrier32_Faults_1" bit 14
   2080: 'Spare_Fault_2080', class No Acknowledgement, trigger "DB302_HMI_Faults_Carrier32_Faults_1" bit 15
   2081: 'Carrier 32 Motion Off Fault', class No Acknowledgement, trigger "DB302_HMI_Faults_Carrier32_Faults_2" bit 0
   2082: 'Carrier 32 Motion On Fault', class No Acknowledgement, trigger "DB302_HMI_Faults_Carrier32_Faults_2" bit 1
   2083: 'Carrier 32 Spacing Fault', class No Acknowledgement, trigger "DB302_HMI_Faults_Carrier32_Faults_2" bit 2
   2084: 'Carrier 32 Duplicate Carrier Number Fault', class No Acknowledgement, trigger "DB302_HMI_Faults_Carrier32_Faults_2" bit 3
   2085: 'Spare_Fault_2085', class No Acknowledgement, trigger "DB302_HMI_Faults_Carrier32_Faults_2" bit 4
   2086: 'Spare_Fault_2086', class No Acknowledgement, trigger "DB302_HMI_Faults_Carrier32_Faults_2" bit 5
   2087: 'Spare_Fault_2087', class No Acknowledgement, trigger "DB302_HMI_Faults_Carrier32_Faults_2" bit 6
   2088: 'Spare_Fault_2088', class No Acknowledgement, trigger "DB302_HMI_Faults_Carrier32_Faults_2" bit 7
   2089: 'Spare_Fault_2089', class No Acknowledgement, trigger "DB302_HMI_Faults_Carrier32_Faults_2" bit 8
   2090: 'Spare_Fault_2090', class No Acknowledgement, trigger "DB302_HMI_Faults_Carrier32_Faults_2" bit 9
   2091: 'Spare_Fault_2091', class No Acknowledgement, trigger "DB302_HMI_Faults_Carrier32_Faults_2" bit 10
   2092: 'Spare_Fault_2092', class No Acknowledgement, trigger "DB302_HMI_Faults_Carrier32_Faults_2" bit 11
   2093: 'Spare_Fault_2093', class No Acknowledgement, trigger "DB302_HMI_Faults_Carrier32_Faults_2" bit 12
   2094: 'Spare_Fault_2094', class No Acknowledgement, trigger "DB302_HMI_Faults_Carrier32_Faults_2" bit 13
   2095: 'Spare_Fault_2095', class No Acknowledgement, trigger "DB302_HMI_Faults_Carrier32_Faults_2" bit 14
   2096: 'Spare_Fault_2096', class No Acknowledgement, trigger "DB302_HMI_Faults_Carrier32_Faults_2" bit 15
   2097: 'Spare_Fault_2097', class No Acknowledgement, trigger "DB302_HMI_Faults_Carrier32_Faults_3" bit 0
   2098: 'Spare_Fault_2098', class No Acknowledgement, trigger "DB302_HMI_Faults_Carrier32_Faults_3" bit 1
   2099: 'Spare_Fault_2099', class No Acknowledgement, trigger "DB302_HMI_Faults_Carrier32_Faults_3" bit 2
   2100: 'Spare_Fault_2100', class No Acknowledgement, trigger "DB302_HMI_Faults_Carrier32_Faults_3" bit 3
   2101: 'Spare_Fault_2101', class No Acknowledgement, trigger "DB302_HMI_Faults_Carrier32_Faults_3" bit 4
   2102: 'Spare_Fault_2102', class No Acknowledgement, trigger "DB302_HMI_Faults_Carrier32_Faults_3" bit 5
   2103: 'Spare_Fault_2103', class No Acknowledgement, trigger "DB302_HMI_Faults_Carrier32_Faults_3" bit 6
   2104: 'Spare_Fault_2104', class No Acknowledgement, trigger "DB302_HMI_Faults_Carrier32_Faults_3" bit 7
   2105: 'Spare_Fault_2105', class No Acknowledgement, trigger "DB302_HMI_Faults_Carrier32_Faults_3" bit 8
   2106: 'Spare_Fault_2106', class No Acknowledgement, trigger "DB302_HMI_Faults_Carrier32_Faults_3" bit 9
   2107: 'Spare_Fault_2107', class No Acknowledgement, trigger "DB302_HMI_Faults_Carrier32_Faults_3" bit 10
   2108: 'Spare_Fault_2108', class No Acknowledgement, trigger "DB302_HMI_Faults_Carrier32_Faults_3" bit 11
   2109: 'Spare_Fault_2109', class No Acknowledgement, trigger "DB302_HMI_Faults_Carrier32_Faults_3" bit 12
   2110: 'Spare_Fault_2110', class No Acknowledgement, trigger "DB302_HMI_Faults_Carrier32_Faults_3" bit 13
   2111: 'Spare_Fault_2111', class No Acknowledgement, trigger "DB302_HMI_Faults_Carrier32_Faults_3" bit 14
   2112: 'Spare_Fault_2112', class No Acknowledgement, trigger "DB302_HMI_Faults_Carrier32_Faults_3" bit 15
   2113: 'Carrier 33 Disconnect Open Power Fault DI11.0', class No Acknowledgement, trigger "DB302_HMI_Faults_Carrier33_Faults_0" bit 0
   2114: 'Carrier 33 Drive Profinet Comm Fault', class No Acknowledgement, trigger "DB302_HMI_Faults_Carrier33_Faults_0" bit 1
   2115: 'Carrier 33 Production Stop Not Reset', class No Acknowledgement, trigger "DB302_HMI_Faults_Carrier33_Faults_0" bit 2
   2116: 'Carrier 33 CB02122 Tripped', class No Acknowledgement, trigger "DB302_HMI_Faults_Carrier33_Faults_0" bit 3
   2117: 'Carrier 33 CB02123 Tripped', class No Acknowledgement, trigger "DB302_HMI_Faults_Carrier33_Faults_0" bit 4
   2118: 'Carrier 33 AUX1 CB Tripped', class No Acknowledgement, trigger "DB302_HMI_Faults_Carrier33_Faults_0" bit 5
   2119: 'Carrier 33 AUX2 CB Tripped', class No Acknowledgement, trigger "DB302_HMI_Faults_Carrier33_Faults_0" bit 6
   2120: 'Carrier 33 PLC Not Communicating', class No Acknowledgement, trigger "DB302_HMI_Faults_Carrier33_Faults_0" bit 7
   2121: 'Carrier 33 Safe Input Card Fault', class No Acknowledgement, trigger "DB302_HMI_Faults_Carrier33_Faults_0" bit 8
   2122: 'Carrier 33 Safe Output Card Fault', class No Acknowledgement, trigger "DB302_HMI_Faults_Carrier33_Faults_0" bit 9
   2123: 'Carrier 33 Standard Input Card Fault', class No Acknowledgement, trigger "DB302_HMI_Faults_Carrier33_Faults_0" bit 10
   2124: 'Carrier 33 Standard Output Card Fault', class No Acknowledgement, trigger "DB302_HMI_Faults_Carrier33_Faults_0" bit 11
   2125: 'Carrier 33 Encoder Position Fault', class No Acknowledgement, trigger "DB302_HMI_Faults_Carrier33_Faults_0" bit 12
   2126: 'Carrier 33 Encoder Internal Error', class No Acknowledgement, trigger "DB302_HMI_Faults_Carrier33_Faults_0" bit 13
   2127: 'Carrier 33 Encoder Comm Fault', class No Acknowledgement, trigger "DB302_HMI_Faults_Carrier33_Faults_0" bit 14
   2128: 'Carrier 33 HMI Comm Fault', class No Acknowledgement, trigger "DB302_HMI_Faults_Carrier33_Faults_0" bit 15
   2129: 'Carrier 33 Crash Detection Fault', class No Acknowledgement, trigger "DB302_HMI_Faults_Carrier33_Faults_1" bit 0
   2130: 'Carrier 33 Carrier Number Invalid', class No Acknowledgement, trigger "DB302_HMI_Faults_Carrier33_Faults_1" bit 1
   2131: 'Carrier 33 Drive: PROFINET configuration error', class No Acknowledgement, trigger "DB302_HMI_Faults_Carrier33_Faults_1" bit 2